DATA_BLOCK "DB_SDC_TS_REFERENCE_3"   // DB3782
{ S7_Optimized_Access := 'FALSE' }
VERSION : 0.1
   VAR
      HEADER : Struct   // Struktur für Datenheader // nicht verschieben
         DB_NR : Int := 3782;   // DB Nummer
         MIN_NR_SEK : Int := 201;   // Niedrigste SEK Nummer im DB
         MAX_NR_SEK : Int := 300;   // Höchste SEK Nummer im DB
         START_DAT : Int := 20;   // Startadresse der SEK im DB
         LAENGE_SEK_DATA : Int := 200;   // Länge SEK Data
         Res10 : Int := 0;   // Reserve
         Res12 : Int := 0;   // Reserve
         Res14 : Int := 0;   // Reserve
         Res16 : Int := 0;   // Reserve
         Res18 : Int := 0;   // Reserve
      END_STRUCT;
      Reference : Array[201..300] of Struct   // Sektionsnummer
         Sektion : Array[1..16] of Char;   // definition Sektion
         Actionpoint_1 : Array[1..16] of Char;   // definition Actionpoint 1
         Actionpoint_2 : Array[1..16] of Char;   // definition Actionpoint 2
         Height : Array[1..16] of Char;   // definition Hubposition (mm)
         Hoist_offset_1 : Array[1..16] of Char;   // definition Hub-Offset 1 (mm)
         Hoist_offset_2 : Array[1..16] of Char;   // definition Hub-Offset 2 (mm)
         Hoist_offset_3 : Array[1..16] of Char;   // definition Hub-Offset 3(mm)
         Hoist_offset_4 : Array[1..16] of Char;   // definition Hub-Offset 4 (mm)
         Reserve : Array[128..199] of Char;
      END_STRUCT;
   END_VAR
BEGIN
   Reference[201].Reserve[199] := ' ';
   Reference[201].Reserve[198] := ' ';
   Reference[201].Reserve[197] := ' ';
   Reference[201].Reserve[196] := ' ';
   Reference[201].Reserve[195] := ' ';
   Reference[201].Reserve[194] := ' ';
   Reference[201].Reserve[193] := ' ';
   Reference[201].Reserve[192] := ' ';
   Reference[201].Reserve[191] := ' ';
   Reference[201].Reserve[190] := ' ';
   Reference[201].Reserve[189] := ' ';
   Reference[201].Reserve[188] := ' ';
   Reference[201].Reserve[187] := ' ';
   Reference[201].Reserve[186] := ' ';
   Reference[201].Reserve[185] := ' ';
   Reference[201].Reserve[184] := ' ';
   Reference[201].Reserve[183] := ' ';
   Reference[201].Reserve[182] := ' ';
   Reference[201].Reserve[181] := ' ';
   Reference[201].Reserve[180] := ' ';
   Reference[201].Reserve[179] := ' ';
   Reference[201].Reserve[178] := ' ';
   Reference[201].Reserve[177] := ' ';
   Reference[201].Reserve[176] := ' ';
   Reference[201].Reserve[175] := ' ';
   Reference[201].Reserve[174] := ' ';
   Reference[201].Reserve[173] := ' ';
   Reference[201].Reserve[172] := ' ';
   Reference[201].Reserve[171] := ' ';
   Reference[201].Reserve[170] := ' ';
   Reference[201].Reserve[169] := ' ';
   Reference[201].Reserve[168] := ' ';
   Reference[201].Reserve[167] := ' ';
   Reference[201].Reserve[166] := ' ';
   Reference[201].Reserve[165] := ' ';
   Reference[201].Reserve[164] := ' ';
   Reference[201].Reserve[163] := ' ';
   Reference[201].Reserve[162] := ' ';
   Reference[201].Reserve[161] := ' ';
   Reference[201].Reserve[160] := ' ';
   Reference[201].Reserve[159] := ' ';
   Reference[201].Reserve[158] := ' ';
   Reference[201].Reserve[157] := ' ';
   Reference[201].Reserve[156] := ' ';
   Reference[201].Reserve[155] := ' ';
   Reference[201].Reserve[154] := ' ';
   Reference[201].Reserve[153] := ' ';
   Reference[201].Reserve[152] := ' ';
   Reference[201].Reserve[151] := ' ';
   Reference[201].Reserve[150] := ' ';
   Reference[201].Reserve[149] := ' ';
   Reference[201].Reserve[148] := ' ';
   Reference[201].Reserve[147] := ' ';
   Reference[201].Reserve[146] := ' ';
   Reference[201].Reserve[145] := ' ';
   Reference[201].Reserve[144] := ' ';
   Reference[201].Reserve[143] := '0';
   Reference[201].Reserve[142] := '0';
   Reference[201].Reserve[141] := '0';
   Reference[201].Reserve[140] := '0';
   Reference[201].Reserve[139] := '0';
   Reference[201].Reserve[138] := '0';
   Reference[201].Reserve[137] := '0';
   Reference[201].Reserve[136] := '0';
   Reference[201].Reserve[135] := '0';
   Reference[201].Reserve[134] := '0';
   Reference[201].Reserve[133] := '0';
   Reference[201].Reserve[132] := '0';
   Reference[201].Reserve[131] := '0';
   Reference[201].Reserve[130] := '0';
   Reference[201].Reserve[129] := '0';
   Reference[201].Reserve[128] := '0';
   Reference[201].Hoist_offset_4[16] := '$00';
   Reference[201].Hoist_offset_4[15] := '$00';
   Reference[201].Hoist_offset_4[14] := '$00';
   Reference[201].Hoist_offset_4[13] := '$00';
   Reference[201].Hoist_offset_4[12] := '$00';
   Reference[201].Hoist_offset_4[11] := '$00';
   Reference[201].Hoist_offset_4[10] := '$00';
   Reference[201].Hoist_offset_4[9] := '$00';
   Reference[201].Hoist_offset_4[8] := '$00';
   Reference[201].Hoist_offset_4[7] := '$00';
   Reference[201].Hoist_offset_4[6] := '$00';
   Reference[201].Hoist_offset_4[5] := '$00';
   Reference[201].Hoist_offset_4[4] := '$00';
   Reference[201].Hoist_offset_4[3] := '$00';
   Reference[201].Hoist_offset_4[2] := '$00';
   Reference[201].Hoist_offset_4[1] := '$00';
   Reference[201].Hoist_offset_3[16] := '$00';
   Reference[201].Hoist_offset_3[15] := '$00';
   Reference[201].Hoist_offset_3[14] := '$00';
   Reference[201].Hoist_offset_3[13] := '$00';
   Reference[201].Hoist_offset_3[12] := '$00';
   Reference[201].Hoist_offset_3[11] := '$00';
   Reference[201].Hoist_offset_3[10] := '$00';
   Reference[201].Hoist_offset_3[9] := '$00';
   Reference[201].Hoist_offset_3[8] := '$00';
   Reference[201].Hoist_offset_3[7] := '$00';
   Reference[201].Hoist_offset_3[6] := '$00';
   Reference[201].Hoist_offset_3[5] := '$00';
   Reference[201].Hoist_offset_3[4] := '$00';
   Reference[201].Hoist_offset_3[3] := '$00';
   Reference[201].Hoist_offset_3[2] := '$00';
   Reference[201].Hoist_offset_3[1] := '$00';
   Reference[201].Hoist_offset_2[16] := '$00';
   Reference[201].Hoist_offset_2[15] := '$00';
   Reference[201].Hoist_offset_2[14] := '$00';
   Reference[201].Hoist_offset_2[13] := '$00';
   Reference[201].Hoist_offset_2[12] := '$00';
   Reference[201].Hoist_offset_2[11] := '$00';
   Reference[201].Hoist_offset_2[10] := '$00';
   Reference[201].Hoist_offset_2[9] := '$00';
   Reference[201].Hoist_offset_2[8] := '$00';
   Reference[201].Hoist_offset_2[7] := '$00';
   Reference[201].Hoist_offset_2[6] := '$00';
   Reference[201].Hoist_offset_2[5] := '$00';
   Reference[201].Hoist_offset_2[4] := '$00';
   Reference[201].Hoist_offset_2[3] := '$00';
   Reference[201].Hoist_offset_2[2] := '$00';
   Reference[201].Hoist_offset_2[1] := '$00';
   Reference[201].Hoist_offset_1[16] := '$00';
   Reference[201].Hoist_offset_1[15] := '$00';
   Reference[201].Hoist_offset_1[14] := '$00';
   Reference[201].Hoist_offset_1[13] := '$00';
   Reference[201].Hoist_offset_1[12] := '$00';
   Reference[201].Hoist_offset_1[11] := '$00';
   Reference[201].Hoist_offset_1[10] := '$00';
   Reference[201].Hoist_offset_1[9] := '$00';
   Reference[201].Hoist_offset_1[8] := '$00';
   Reference[201].Hoist_offset_1[7] := '$00';
   Reference[201].Hoist_offset_1[6] := '$00';
   Reference[201].Hoist_offset_1[5] := '$00';
   Reference[201].Hoist_offset_1[4] := '$00';
   Reference[201].Hoist_offset_1[3] := '$00';
   Reference[201].Hoist_offset_1[2] := '$00';
   Reference[201].Hoist_offset_1[1] := '$00';
   Reference[201].Height[16] := '$00';
   Reference[201].Height[15] := '$00';
   Reference[201].Height[14] := '$00';
   Reference[201].Height[13] := '$00';
   Reference[201].Height[12] := '$00';
   Reference[201].Height[11] := '$00';
   Reference[201].Height[10] := '$00';
   Reference[201].Height[9] := '$00';
   Reference[201].Height[8] := '$00';
   Reference[201].Height[7] := '$00';
   Reference[201].Height[6] := '$00';
   Reference[201].Height[5] := '$00';
   Reference[201].Height[4] := '$00';
   Reference[201].Height[3] := '$00';
   Reference[201].Height[2] := '$00';
   Reference[201].Height[1] := '$00';
   Reference[201].Actionpoint_2[16] := '0';
   Reference[201].Actionpoint_2[15] := '0';
   Reference[201].Actionpoint_2[14] := '0';
   Reference[201].Actionpoint_2[13] := '0';
   Reference[201].Actionpoint_2[12] := '0';
   Reference[201].Actionpoint_2[11] := '0';
   Reference[201].Actionpoint_2[10] := '0';
   Reference[201].Actionpoint_2[9] := '0';
   Reference[201].Actionpoint_2[8] := '0';
   Reference[201].Actionpoint_2[7] := '0';
   Reference[201].Actionpoint_2[6] := '0';
   Reference[201].Actionpoint_2[5] := '0';
   Reference[201].Actionpoint_2[4] := '0';
   Reference[201].Actionpoint_2[3] := '0';
   Reference[201].Actionpoint_2[2] := '0';
   Reference[201].Actionpoint_2[1] := '0';
   Reference[201].Actionpoint_1[16] := '0';
   Reference[201].Actionpoint_1[15] := '0';
   Reference[201].Actionpoint_1[14] := '0';
   Reference[201].Actionpoint_1[13] := '0';
   Reference[201].Actionpoint_1[12] := '0';
   Reference[201].Actionpoint_1[11] := '0';
   Reference[201].Actionpoint_1[10] := '0';
   Reference[201].Actionpoint_1[9] := '0';
   Reference[201].Actionpoint_1[8] := '0';
   Reference[201].Actionpoint_1[7] := '0';
   Reference[201].Actionpoint_1[6] := '0';
   Reference[201].Actionpoint_1[5] := '0';
   Reference[201].Actionpoint_1[4] := '0';
   Reference[201].Actionpoint_1[3] := '0';
   Reference[201].Actionpoint_1[2] := '0';
   Reference[201].Actionpoint_1[1] := '0';
   Reference[201].Sektion[1] := ' ';
   Reference[201].Sektion[2] := ' ';
   Reference[201].Sektion[3] := ' ';
   Reference[201].Sektion[4] := ' ';
   Reference[201].Sektion[5] := ' ';
   Reference[201].Sektion[6] := ' ';
   Reference[201].Sektion[7] := ' ';
   Reference[201].Sektion[8] := ' ';
   Reference[201].Sektion[9] := ' ';
   Reference[201].Sektion[10] := ' ';
   Reference[201].Sektion[11] := ' ';
   Reference[201].Sektion[12] := ' ';
   Reference[201].Sektion[13] := ' ';
   Reference[201].Sektion[14] := ' ';
   Reference[201].Sektion[15] := ' ';
   Reference[201].Sektion[16] := ' ';
   // 19800 more start values not shown
END_DATA_BLOCK

DATA_BLOCK "DB_SDC_TS_REFERENCE_4"   // DB3783
{ S7_Optimized_Access := 'FALSE' }
VERSION : 0.1
   VAR
      HEADER : Struct   // Struktur für Datenheader // nicht verschieben
         DB_NR : Int := 3783;   // DB Nummer
         MIN_NR_SEK : Int := 301;   // Niedrigste SEK Nummer im DB
         MAX_NR_SEK : Int := 400;   // Höchste SEK Nummer im DB
         START_DAT : Int := 20;   // Startadresse der SEK im DB
         LAENGE_SEK_DATA : Int := 200;   // Länge SEK Data
         Res10 : Int := 0;   // Reserve
         Res12 : Int := 0;   // Reserve
         Res14 : Int := 0;   // Reserve
         Res16 : Int := 0;   // Reserve
         Res18 : Int := 0;   // Reserve
      END_STRUCT;
      Reference : Array[301..400] of Struct   // Sektionsnummer
         Sektion : Array[1..16] of Char;   // definition Sektion
         Actionpoint_1 : Array[1..16] of Char;   // definition Actionpoint 1
         Actionpoint_2 : Array[1..16] of Char;   // definition Actionpoint 2
         Height : Array[1..16] of Char;   // definition Hubposition (mm)
         Hoist_offset_1 : Array[1..16] of Char;   // definition Hub-Offset 1 (mm)
         Hoist_offset_2 : Array[1..16] of Char;   // definition Hub-Offset 2 (mm)
         Hoist_offset_3 : Array[1..16] of Char;   // definition Hub-Offset 3(mm)
         Hoist_offset_4 : Array[1..16] of Char;   // definition Hub-Offset 4 (mm)
         Reserve : Array[128..199] of Char;
      END_STRUCT;
   END_VAR
BEGIN
   Reference[301].Reserve[199] := ' ';
   Reference[301].Reserve[198] := ' ';
   Reference[301].Reserve[197] := ' ';
   Reference[301].Reserve[196] := ' ';
   Reference[301].Reserve[195] := ' ';
   Reference[301].Reserve[194] := ' ';
   Reference[301].Reserve[193] := ' ';
   Reference[301].Reserve[192] := ' ';
   Reference[301].Reserve[191] := ' ';
   Reference[301].Reserve[190] := ' ';
   Reference[301].Reserve[189] := ' ';
   Reference[301].Reserve[188] := ' ';
   Reference[301].Reserve[187] := ' ';
   Reference[301].Reserve[186] := ' ';
   Reference[301].Reserve[185] := ' ';
   Reference[301].Reserve[184] := ' ';
   Reference[301].Reserve[183] := ' ';
   Reference[301].Reserve[182] := ' ';
   Reference[301].Reserve[181] := ' ';
   Reference[301].Reserve[180] := ' ';
   Reference[301].Reserve[179] := ' ';
   Reference[301].Reserve[178] := ' ';
   Reference[301].Reserve[177] := ' ';
   Reference[301].Reserve[176] := ' ';
   Reference[301].Reserve[175] := ' ';
   Reference[301].Reserve[174] := ' ';
   Reference[301].Reserve[173] := ' ';
   Reference[301].Reserve[172] := ' ';
   Reference[301].Reserve[171] := ' ';
   Reference[301].Reserve[170] := ' ';
   Reference[301].Reserve[169] := ' ';
   Reference[301].Reserve[168] := ' ';
   Reference[301].Reserve[167] := ' ';
   Reference[301].Reserve[166] := ' ';
   Reference[301].Reserve[165] := ' ';
   Reference[301].Reserve[164] := ' ';
   Reference[301].Reserve[163] := ' ';
   Reference[301].Reserve[162] := ' ';
   Reference[301].Reserve[161] := ' ';
   Reference[301].Reserve[160] := ' ';
   Reference[301].Reserve[159] := ' ';
   Reference[301].Reserve[158] := ' ';
   Reference[301].Reserve[157] := ' ';
   Reference[301].Reserve[156] := ' ';
   Reference[301].Reserve[155] := ' ';
   Reference[301].Reserve[154] := ' ';
   Reference[301].Reserve[153] := ' ';
   Reference[301].Reserve[152] := ' ';
   Reference[301].Reserve[151] := ' ';
   Reference[301].Reserve[150] := ' ';
   Reference[301].Reserve[149] := ' ';
   Reference[301].Reserve[148] := ' ';
   Reference[301].Reserve[147] := ' ';
   Reference[301].Reserve[146] := ' ';
   Reference[301].Reserve[145] := ' ';
   Reference[301].Reserve[144] := ' ';
   Reference[301].Reserve[143] := '0';
   Reference[301].Reserve[142] := '0';
   Reference[301].Reserve[141] := '0';
   Reference[301].Reserve[140] := '0';
   Reference[301].Reserve[139] := '0';
   Reference[301].Reserve[138] := '0';
   Reference[301].Reserve[137] := '0';
   Reference[301].Reserve[136] := '0';
   Reference[301].Reserve[135] := '0';
   Reference[301].Reserve[134] := '0';
   Reference[301].Reserve[133] := '0';
   Reference[301].Reserve[132] := '0';
   Reference[301].Reserve[131] := '0';
   Reference[301].Reserve[130] := '0';
   Reference[301].Reserve[129] := '0';
   Reference[301].Reserve[128] := '0';
   Reference[301].Hoist_offset_4[16] := '$00';
   Reference[301].Hoist_offset_4[15] := '$00';
   Reference[301].Hoist_offset_4[14] := '$00';
   Reference[301].Hoist_offset_4[13] := '$00';
   Reference[301].Hoist_offset_4[12] := '$00';
   Reference[301].Hoist_offset_4[11] := '$00';
   Reference[301].Hoist_offset_4[10] := '$00';
   Reference[301].Hoist_offset_4[9] := '$00';
   Reference[301].Hoist_offset_4[8] := '$00';
   Reference[301].Hoist_offset_4[7] := '$00';
   Reference[301].Hoist_offset_4[6] := '$00';
   Reference[301].Hoist_offset_4[5] := '$00';
   Reference[301].Hoist_offset_4[4] := '$00';
   Reference[301].Hoist_offset_4[3] := '$00';
   Reference[301].Hoist_offset_4[2] := '$00';
   Reference[301].Hoist_offset_4[1] := '$00';
   Reference[301].Hoist_offset_3[16] := '$00';
   Reference[301].Hoist_offset_3[15] := '$00';
   Reference[301].Hoist_offset_3[14] := '$00';
   Reference[301].Hoist_offset_3[13] := '$00';
   Reference[301].Hoist_offset_3[12] := '$00';
   Reference[301].Hoist_offset_3[11] := '$00';
   Reference[301].Hoist_offset_3[10] := '$00';
   Reference[301].Hoist_offset_3[9] := '$00';
   Reference[301].Hoist_offset_3[8] := '$00';
   Reference[301].Hoist_offset_3[7] := '$00';
   Reference[301].Hoist_offset_3[6] := '$00';
   Reference[301].Hoist_offset_3[5] := '$00';
   Reference[301].Hoist_offset_3[4] := '$00';
   Reference[301].Hoist_offset_3[3] := '$00';
   Reference[301].Hoist_offset_3[2] := '$00';
   Reference[301].Hoist_offset_3[1] := '$00';
   Reference[301].Hoist_offset_2[16] := '$00';
   Reference[301].Hoist_offset_2[15] := '$00';
   Reference[301].Hoist_offset_2[14] := '$00';
   Reference[301].Hoist_offset_2[13] := '$00';
   Reference[301].Hoist_offset_2[12] := '$00';
   Reference[301].Hoist_offset_2[11] := '$00';
   Reference[301].Hoist_offset_2[10] := '$00';
   Reference[301].Hoist_offset_2[9] := '$00';
   Reference[301].Hoist_offset_2[8] := '$00';
   Reference[301].Hoist_offset_2[7] := '$00';
   Reference[301].Hoist_offset_2[6] := '$00';
   Reference[301].Hoist_offset_2[5] := '$00';
   Reference[301].Hoist_offset_2[4] := '$00';
   Reference[301].Hoist_offset_2[3] := '$00';
   Reference[301].Hoist_offset_2[2] := '$00';
   Reference[301].Hoist_offset_2[1] := '$00';
   Reference[301].Hoist_offset_1[16] := '$00';
   Reference[301].Hoist_offset_1[15] := '$00';
   Reference[301].Hoist_offset_1[14] := '$00';
   Reference[301].Hoist_offset_1[13] := '$00';
   Reference[301].Hoist_offset_1[12] := '$00';
   Reference[301].Hoist_offset_1[11] := '$00';
   Reference[301].Hoist_offset_1[10] := '$00';
   Reference[301].Hoist_offset_1[9] := '$00';
   Reference[301].Hoist_offset_1[8] := '$00';
   Reference[301].Hoist_offset_1[7] := '$00';
   Reference[301].Hoist_offset_1[6] := '$00';
   Reference[301].Hoist_offset_1[5] := '$00';
   Reference[301].Hoist_offset_1[4] := '$00';
   Reference[301].Hoist_offset_1[3] := '$00';
   Reference[301].Hoist_offset_1[2] := '$00';
   Reference[301].Hoist_offset_1[1] := '$00';
   Reference[301].Height[16] := '$00';
   Reference[301].Height[15] := '$00';
   Reference[301].Height[14] := '$00';
   Reference[301].Height[13] := '$00';
   Reference[301].Height[12] := '$00';
   Reference[301].Height[11] := '$00';
   Reference[301].Height[10] := '$00';
   Reference[301].Height[9] := '$00';
   Reference[301].Height[8] := '$00';
   Reference[301].Height[7] := '$00';
   Reference[301].Height[6] := '$00';
   Reference[301].Height[5] := '$00';
   Reference[301].Height[4] := '$00';
   Reference[301].Height[3] := '$00';
   Reference[301].Height[2] := '$00';
   Reference[301].Height[1] := '$00';
   Reference[301].Actionpoint_2[16] := '0';
   Reference[301].Actionpoint_2[15] := '0';
   Reference[301].Actionpoint_2[14] := '0';
   Reference[301].Actionpoint_2[13] := '0';
   Reference[301].Actionpoint_2[12] := '0';
   Reference[301].Actionpoint_2[11] := '0';
   Reference[301].Actionpoint_2[10] := '0';
   Reference[301].Actionpoint_2[9] := '0';
   Reference[301].Actionpoint_2[8] := '0';
   Reference[301].Actionpoint_2[7] := '0';
   Reference[301].Actionpoint_2[6] := '0';
   Reference[301].Actionpoint_2[5] := '0';
   Reference[301].Actionpoint_2[4] := '0';
   Reference[301].Actionpoint_2[3] := '0';
   Reference[301].Actionpoint_2[2] := '0';
   Reference[301].Actionpoint_2[1] := '0';
   Reference[301].Actionpoint_1[16] := '0';
   Reference[301].Actionpoint_1[15] := '0';
   Reference[301].Actionpoint_1[14] := '0';
   Reference[301].Actionpoint_1[13] := '0';
   Reference[301].Actionpoint_1[12] := '0';
   Reference[301].Actionpoint_1[11] := '0';
   Reference[301].Actionpoint_1[10] := '0';
   Reference[301].Actionpoint_1[9] := '0';
   Reference[301].Actionpoint_1[8] := '0';
   Reference[301].Actionpoint_1[7] := '0';
   Reference[301].Actionpoint_1[6] := '0';
   Reference[301].Actionpoint_1[5] := '0';
   Reference[301].Actionpoint_1[4] := '0';
   Reference[301].Actionpoint_1[3] := '0';
   Reference[301].Actionpoint_1[2] := '0';
   Reference[301].Actionpoint_1[1] := '0';
   Reference[301].Sektion[1] := ' ';
   Reference[301].Sektion[2] := ' ';
   Reference[301].Sektion[3] := ' ';
   Reference[301].Sektion[4] := ' ';
   Reference[301].Sektion[5] := ' ';
   Reference[301].Sektion[6] := ' ';
   Reference[301].Sektion[7] := ' ';
   Reference[301].Sektion[8] := ' ';
   Reference[301].Sektion[9] := ' ';
   Reference[301].Sektion[10] := ' ';
   Reference[301].Sektion[11] := ' ';
   Reference[301].Sektion[12] := ' ';
   Reference[301].Sektion[13] := ' ';
   Reference[301].Sektion[14] := ' ';
   Reference[301].Sektion[15] := ' ';
   Reference[301].Sektion[16] := ' ';
   // 19800 more start values not shown
END_DATA_BLOCK

DATA_BLOCK "DB_SDC_TS_REFERENCE_5"   // DB3784
{ S7_Optimized_Access := 'FALSE' }
VERSION : 0.1
   VAR
      HEADER : Struct   // Struktur für Datenheader // nicht verschieben
         DB_NR : Int := 3784;   // DB Nummer
         MIN_NR_SEK : Int := 401;   // Niedrigste SEK Nummer im DB
         MAX_NR_SEK : Int := 500;   // Höchste SEK Nummer im DB
         START_DAT : Int := 20;   // Startadresse der SEK im DB
         LAENGE_SEK_DATA : Int := 200;   // Länge SEK Data
         Res10 : Int := 0;   // Reserve
         Res12 : Int := 0;   // Reserve
         Res14 : Int := 0;   // Reserve
         Res16 : Int := 0;   // Reserve
         Res18 : Int := 0;   // Reserve
      END_STRUCT;
      Reference : Array[401..500] of Struct   // Sektionsnummer
         Sektion : Array[1..16] of Char;   // definition Sektion
         Actionpoint_1 : Array[1..16] of Char;   // definition Actionpoint 1
         Actionpoint_2 : Array[1..16] of Char;   // definition Actionpoint 2
         Height : Array[1..16] of Char;   // definition Hubposition (mm)
         Hoist_offset_1 : Array[1..16] of Char;   // definition Hub-Offset 1 (mm)
         Hoist_offset_2 : Array[1..16] of Char;   // definition Hub-Offset 2 (mm)
         Hoist_offset_3 : Array[1..16] of Char;   // definition Hub-Offset 3(mm)
         Hoist_offset_4 : Array[1..16] of Char;   // definition Hub-Offset 4 (mm)
         Reserve : Array[128..199] of Char;
      END_STRUCT;
   END_VAR
BEGIN
   Reference[401].Reserve[199] := ' ';
   Reference[401].Reserve[198] := ' ';
   Reference[401].Reserve[197] := ' ';
   Reference[401].Reserve[196] := ' ';
   Reference[401].Reserve[195] := ' ';
   Reference[401].Reserve[194] := ' ';
   Reference[401].Reserve[193] := ' ';
   Reference[401].Reserve[192] := ' ';
   Reference[401].Reserve[191] := ' ';
   Reference[401].Reserve[190] := ' ';
   Reference[401].Reserve[189] := ' ';
   Reference[401].Reserve[188] := ' ';
   Reference[401].Reserve[187] := ' ';
   Reference[401].Reserve[186] := ' ';
   Reference[401].Reserve[185] := ' ';
   Reference[401].Reserve[184] := ' ';
   Reference[401].Reserve[183] := ' ';
   Reference[401].Reserve[182] := ' ';
   Reference[401].Reserve[181] := ' ';
   Reference[401].Reserve[180] := ' ';
   Reference[401].Reserve[179] := ' ';
   Reference[401].Reserve[178] := ' ';
   Reference[401].Reserve[177] := ' ';
   Reference[401].Reserve[176] := ' ';
   Reference[401].Reserve[175] := ' ';
   Reference[401].Reserve[174] := ' ';
   Reference[401].Reserve[173] := ' ';
   Reference[401].Reserve[172] := ' ';
   Reference[401].Reserve[171] := ' ';
   Reference[401].Reserve[170] := ' ';
   Reference[401].Reserve[169] := ' ';
   Reference[401].Reserve[168] := ' ';
   Reference[401].Reserve[167] := ' ';
   Reference[401].Reserve[166] := ' ';
   Reference[401].Reserve[165] := ' ';
   Reference[401].Reserve[164] := ' ';
   Reference[401].Reserve[163] := ' ';
   Reference[401].Reserve[162] := ' ';
   Reference[401].Reserve[161] := ' ';
   Reference[401].Reserve[160] := ' ';
   Reference[401].Reserve[159] := ' ';
   Reference[401].Reserve[158] := ' ';
   Reference[401].Reserve[157] := ' ';
   Reference[401].Reserve[156] := ' ';
   Reference[401].Reserve[155] := ' ';
   Reference[401].Reserve[154] := ' ';
   Reference[401].Reserve[153] := ' ';
   Reference[401].Reserve[152] := ' ';
   Reference[401].Reserve[151] := ' ';
   Reference[401].Reserve[150] := ' ';
   Reference[401].Reserve[149] := ' ';
   Reference[401].Reserve[148] := ' ';
   Reference[401].Reserve[147] := ' ';
   Reference[401].Reserve[146] := ' ';
   Reference[401].Reserve[145] := ' ';
   Reference[401].Reserve[144] := ' ';
   Reference[401].Reserve[143] := '0';
   Reference[401].Reserve[142] := '0';
   Reference[401].Reserve[141] := '0';
   Reference[401].Reserve[140] := '0';
   Reference[401].Reserve[139] := '0';
   Reference[401].Reserve[138] := '0';
   Reference[401].Reserve[137] := '0';
   Reference[401].Reserve[136] := '0';
   Reference[401].Reserve[135] := '0';
   Reference[401].Reserve[134] := '0';
   Reference[401].Reserve[133] := '0';
   Reference[401].Reserve[132] := '0';
   Reference[401].Reserve[131] := '0';
   Reference[401].Reserve[130] := '0';
   Reference[401].Reserve[129] := '0';
   Reference[401].Reserve[128] := '0';
   Reference[401].Hoist_offset_4[16] := '$00';
   Reference[401].Hoist_offset_4[15] := '$00';
   Reference[401].Hoist_offset_4[14] := '$00';
   Reference[401].Hoist_offset_4[13] := '$00';
   Reference[401].Hoist_offset_4[12] := '$00';
   Reference[401].Hoist_offset_4[11] := '$00';
   Reference[401].Hoist_offset_4[10] := '$00';
   Reference[401].Hoist_offset_4[9] := '$00';
   Reference[401].Hoist_offset_4[8] := '$00';
   Reference[401].Hoist_offset_4[7] := '$00';
   Reference[401].Hoist_offset_4[6] := '$00';
   Reference[401].Hoist_offset_4[5] := '$00';
   Reference[401].Hoist_offset_4[4] := '$00';
   Reference[401].Hoist_offset_4[3] := '$00';
   Reference[401].Hoist_offset_4[2] := '$00';
   Reference[401].Hoist_offset_4[1] := '$00';
   Reference[401].Hoist_offset_3[16] := '$00';
   Reference[401].Hoist_offset_3[15] := '$00';
   Reference[401].Hoist_offset_3[14] := '$00';
   Reference[401].Hoist_offset_3[13] := '$00';
   Reference[401].Hoist_offset_3[12] := '$00';
   Reference[401].Hoist_offset_3[11] := '$00';
   Reference[401].Hoist_offset_3[10] := '$00';
   Reference[401].Hoist_offset_3[9] := '$00';
   Reference[401].Hoist_offset_3[8] := '$00';
   Reference[401].Hoist_offset_3[7] := '$00';
   Reference[401].Hoist_offset_3[6] := '$00';
   Reference[401].Hoist_offset_3[5] := '$00';
   Reference[401].Hoist_offset_3[4] := '$00';
   Reference[401].Hoist_offset_3[3] := '$00';
   Reference[401].Hoist_offset_3[2] := '$00';
   Reference[401].Hoist_offset_3[1] := '$00';
   Reference[401].Hoist_offset_2[16] := '$00';
   Reference[401].Hoist_offset_2[15] := '$00';
   Reference[401].Hoist_offset_2[14] := '$00';
   Reference[401].Hoist_offset_2[13] := '$00';
   Reference[401].Hoist_offset_2[12] := '$00';
   Reference[401].Hoist_offset_2[11] := '$00';
   Reference[401].Hoist_offset_2[10] := '$00';
   Reference[401].Hoist_offset_2[9] := '$00';
   Reference[401].Hoist_offset_2[8] := '$00';
   Reference[401].Hoist_offset_2[7] := '$00';
   Reference[401].Hoist_offset_2[6] := '$00';
   Reference[401].Hoist_offset_2[5] := '$00';
   Reference[401].Hoist_offset_2[4] := '$00';
   Reference[401].Hoist_offset_2[3] := '$00';
   Reference[401].Hoist_offset_2[2] := '$00';
   Reference[401].Hoist_offset_2[1] := '$00';
   Reference[401].Hoist_offset_1[16] := '$00';
   Reference[401].Hoist_offset_1[15] := '$00';
   Reference[401].Hoist_offset_1[14] := '$00';
   Reference[401].Hoist_offset_1[13] := '$00';
   Reference[401].Hoist_offset_1[12] := '$00';
   Reference[401].Hoist_offset_1[11] := '$00';
   Reference[401].Hoist_offset_1[10] := '$00';
   Reference[401].Hoist_offset_1[9] := '$00';
   Reference[401].Hoist_offset_1[8] := '$00';
   Reference[401].Hoist_offset_1[7] := '$00';
   Reference[401].Hoist_offset_1[6] := '$00';
   Reference[401].Hoist_offset_1[5] := '$00';
   Reference[401].Hoist_offset_1[4] := '$00';
   Reference[401].Hoist_offset_1[3] := '$00';
   Reference[401].Hoist_offset_1[2] := '$00';
   Reference[401].Hoist_offset_1[1] := '$00';
   Reference[401].Height[16] := '$00';
   Reference[401].Height[15] := '$00';
   Reference[401].Height[14] := '$00';
   Reference[401].Height[13] := '$00';
   Reference[401].Height[12] := '$00';
   Reference[401].Height[11] := '$00';
   Reference[401].Height[10] := '$00';
   Reference[401].Height[9] := '$00';
   Reference[401].Height[8] := '$00';
   Reference[401].Height[7] := '$00';
   Reference[401].Height[6] := '$00';
   Reference[401].Height[5] := '$00';
   Reference[401].Height[4] := '$00';
   Reference[401].Height[3] := '$00';
   Reference[401].Height[2] := '$00';
   Reference[401].Height[1] := '$00';
   Reference[401].Actionpoint_2[16] := '0';
   Reference[401].Actionpoint_2[15] := '0';
   Reference[401].Actionpoint_2[14] := '0';
   Reference[401].Actionpoint_2[13] := '0';
   Reference[401].Actionpoint_2[12] := '0';
   Reference[401].Actionpoint_2[11] := '0';
   Reference[401].Actionpoint_2[10] := '0';
   Reference[401].Actionpoint_2[9] := '0';
   Reference[401].Actionpoint_2[8] := '0';
   Reference[401].Actionpoint_2[7] := '0';
   Reference[401].Actionpoint_2[6] := '0';
   Reference[401].Actionpoint_2[5] := '0';
   Reference[401].Actionpoint_2[4] := '0';
   Reference[401].Actionpoint_2[3] := '0';
   Reference[401].Actionpoint_2[2] := '0';
   Reference[401].Actionpoint_2[1] := '0';
   Reference[401].Actionpoint_1[16] := '0';
   Reference[401].Actionpoint_1[15] := '0';
   Reference[401].Actionpoint_1[14] := '0';
   Reference[401].Actionpoint_1[13] := '0';
   Reference[401].Actionpoint_1[12] := '0';
   Reference[401].Actionpoint_1[11] := '0';
   Reference[401].Actionpoint_1[10] := '0';
   Reference[401].Actionpoint_1[9] := '0';
   Reference[401].Actionpoint_1[8] := '0';
   Reference[401].Actionpoint_1[7] := '0';
   Reference[401].Actionpoint_1[6] := '0';
   Reference[401].Actionpoint_1[5] := '0';
   Reference[401].Actionpoint_1[4] := '0';
   Reference[401].Actionpoint_1[3] := '0';
   Reference[401].Actionpoint_1[2] := '0';
   Reference[401].Actionpoint_1[1] := '0';
   Reference[401].Sektion[1] := 'b';
   Reference[401].Sektion[2] := 'u';
   Reference[401].Sektion[3] := 'f';
   Reference[401].Sektion[4] := 'f';
   Reference[401].Sektion[5] := 'e';
   Reference[401].Sektion[6] := 'r';
   Reference[401].Sektion[7] := '$00';
   Reference[401].Sektion[8] := '$00';
   Reference[401].Sektion[9] := '$00';
   Reference[401].Sektion[10] := '$00';
   Reference[401].Sektion[11] := '$00';
   Reference[401].Sektion[12] := '$00';
   Reference[401].Sektion[13] := '$00';
   Reference[401].Sektion[14] := '$00';
   Reference[401].Sektion[15] := '$00';
   Reference[401].Sektion[16] := '$00';
   // 19800 more start values not shown
END_DATA_BLOCK

DATA_BLOCK "DB_SDC_TS_REFERENCE_6"   // DB3785
{ S7_Optimized_Access := 'FALSE' }
VERSION : 0.1
   VAR
      HEADER : Struct   // Struktur für Datenheader // nicht verschieben
         DB_NR : Int := 3785;   // DB Nummer
         MIN_NR_SEK : Int := 501;   // Niedrigste SEK Nummer im DB
         MAX_NR_SEK : Int := 600;   // Höchste SEK Nummer im DB
         START_DAT : Int := 20;   // Startadresse der SEK im DB
         LAENGE_SEK_DATA : Int := 200;   // Länge SEK Data
         Res10 : Int := 0;   // Reserve
         Res12 : Int := 0;   // Reserve
         Res14 : Int := 0;   // Reserve
         Res16 : Int := 0;   // Reserve
         Res18 : Int := 0;   // Reserve
      END_STRUCT;
      Reference : Array[501..600] of Struct   // Sektionsnummer
         Sektion : Array[1..16] of Char;   // definition Sektion
         Actionpoint_1 : Array[1..16] of Char;   // definition Actionpoint 1
         Actionpoint_2 : Array[1..16] of Char;   // definition Actionpoint 2
         Height : Array[1..16] of Char;   // definition Hubposition (mm)
         Hoist_offset_1 : Array[1..16] of Char;   // definition Hub-Offset 1 (mm)
         Hoist_offset_2 : Array[1..16] of Char;   // definition Hub-Offset 2 (mm)
         Hoist_offset_3 : Array[1..16] of Char;   // definition Hub-Offset 3(mm)
         Hoist_offset_4 : Array[1..16] of Char;   // definition Hub-Offset 4 (mm)
         Reserve : Array[128..199] of Char;
      END_STRUCT;
   END_VAR
BEGIN
   Reference[501].Reserve[199] := ' ';
   Reference[501].Reserve[198] := ' ';
   Reference[501].Reserve[197] := ' ';
   Reference[501].Reserve[196] := ' ';
   Reference[501].Reserve[195] := ' ';
   Reference[501].Reserve[194] := ' ';
   Reference[501].Reserve[193] := ' ';
   Reference[501].Reserve[192] := ' ';
   Reference[501].Reserve[191] := ' ';
   Reference[501].Reserve[190] := ' ';
   Reference[501].Reserve[189] := ' ';
   Reference[501].Reserve[188] := ' ';
   Reference[501].Reserve[187] := ' ';
   Reference[501].Reserve[186] := ' ';
   Reference[501].Reserve[185] := ' ';
   Reference[501].Reserve[184] := ' ';
   Reference[501].Reserve[183] := ' ';
   Reference[501].Reserve[182] := ' ';
   Reference[501].Reserve[181] := ' ';
   Reference[501].Reserve[180] := ' ';
   Reference[501].Reserve[179] := ' ';
   Reference[501].Reserve[178] := ' ';
   Reference[501].Reserve[177] := ' ';
   Reference[501].Reserve[176] := ' ';
   Reference[501].Reserve[175] := ' ';
   Reference[501].Reserve[174] := ' ';
   Reference[501].Reserve[173] := ' ';
   Reference[501].Reserve[172] := ' ';
   Reference[501].Reserve[171] := ' ';
   Reference[501].Reserve[170] := ' ';
   Reference[501].Reserve[169] := ' ';
   Reference[501].Reserve[168] := ' ';
   Reference[501].Reserve[167] := ' ';
   Reference[501].Reserve[166] := ' ';
   Reference[501].Reserve[165] := ' ';
   Reference[501].Reserve[164] := ' ';
   Reference[501].Reserve[163] := ' ';
   Reference[501].Reserve[162] := ' ';
   Reference[501].Reserve[161] := ' ';
   Reference[501].Reserve[160] := ' ';
   Reference[501].Reserve[159] := ' ';
   Reference[501].Reserve[158] := ' ';
   Reference[501].Reserve[157] := ' ';
   Reference[501].Reserve[156] := ' ';
   Reference[501].Reserve[155] := ' ';
   Reference[501].Reserve[154] := ' ';
   Reference[501].Reserve[153] := ' ';
   Reference[501].Reserve[152] := ' ';
   Reference[501].Reserve[151] := ' ';
   Reference[501].Reserve[150] := ' ';
   Reference[501].Reserve[149] := ' ';
   Reference[501].Reserve[148] := ' ';
   Reference[501].Reserve[147] := ' ';
   Reference[501].Reserve[146] := ' ';
   Reference[501].Reserve[145] := ' ';